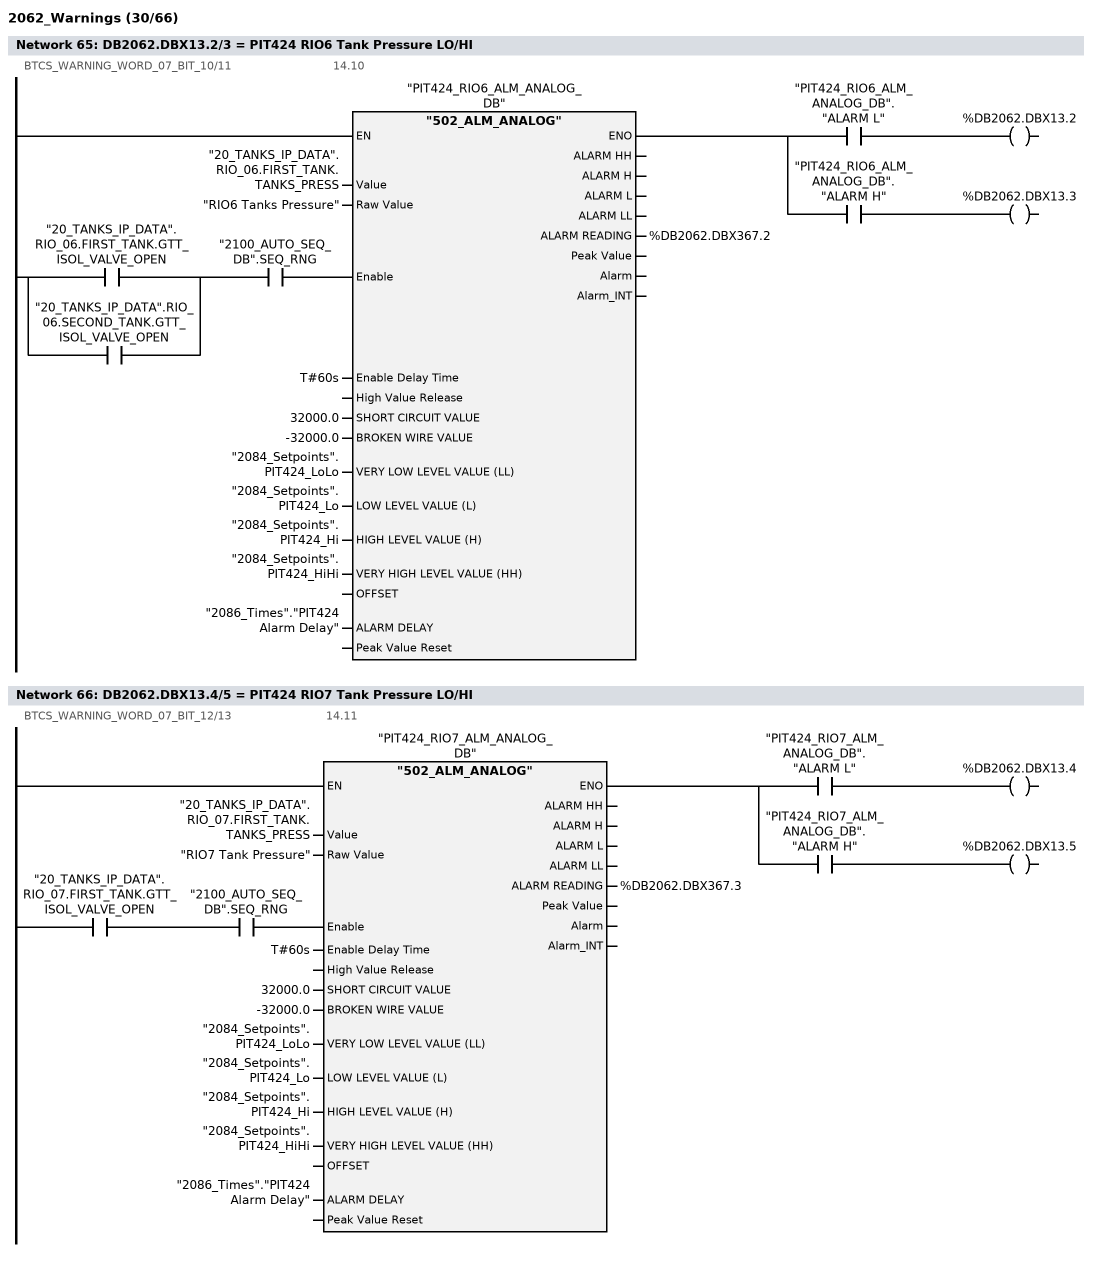
   RUNG wire#powerrail
      "PIT424_RIO6_ALM_ANALOG_DB"(Enable := wire#w2, Value := "20_TANKS_IP_DATA".RIO_06.FIRST_TANK.TANKS_PRESS, "Raw Value" := "RIO6 Tanks Pressure", "Enable Delay Time" := T#60s, "High Value Release" :=, "SHORT CIRCUIT VALUE" := 32000.0, "BROKEN WIRE VALUE" := -32000.0, "VERY LOW LEVEL VALUE (LL)" := "2084_Setpoints".PIT424_LoLo, "LOW LEVEL VALUE (L)" := "2084_Setpoints".PIT424_Lo, "HIGH LEVEL VALUE (H)" := "2084_Setpoints".PIT424_Hi, "VERY HIGH LEVEL VALUE (HH)" := "2084_Setpoints".PIT424_HiHi, OFFSET :=, "ALARM DELAY" := "2086_Times"."PIT424 Alarm Delay", "Peak Value Reset" :=, "ALARM HH" =>, "ALARM H" =>, "ALARM L" =>, "ALARM LL" =>, "ALARM READING" => %DB2062.DBX367.2, "Peak Value" =>, Alarm =>, Alarm_INT =>)
      wire#w3
      Contact( "PIT424_RIO6_ALM_ANALOG_DB"."ALARM L" )
      Coil( %DB2062.DBX13.2 )
   END_RUNG
   RUNG wire#powerrail
      Contact( "20_TANKS_IP_DATA".RIO_06.FIRST_TANK.GTT_ISOL_VALVE_OPEN )
      wire#w1
      Contact( "2100_AUTO_SEQ_DB".SEQ_RNG )
   END_RUNG wire#w2
   RUNG wire#powerrail
      Contact( "20_TANKS_IP_DATA".RIO_06.SECOND_TANK.GTT_ISOL_VALVE_OPEN )
   END_RUNG wire#w1
   RUNG wire#w3
      Contact( "PIT424_RIO6_ALM_ANALOG_DB"."ALARM H" )
      Coil( %DB2062.DBX13.3 )
   END_RUNG
   // the same network as SCL:
   "PIT424_RIO6_ALM_ANALOG_DB"(Value := "20_TANKS_IP_DATA".RIO_06.FIRST_TANK.TANKS_PRESS,   // "502_ALM_ANALOG"
                           "Raw Value" := "RIO6 Tanks Pressure",
                           Enable := ("20_TANKS_IP_DATA".RIO_06.FIRST_TANK.GTT_ISOL_VALVE_OPEN OR "20_TANKS_IP_DATA".RIO_06.SECOND_TANK.GTT_ISOL_VALVE_OPEN) AND "2100_AUTO_SEQ_DB".SEQ_RNG,
                           "Enable Delay Time" := T#60s,
                           "SHORT CIRCUIT VALUE" := 32000.0,
                           "BROKEN WIRE VALUE" := -32000.0,
                           "VERY LOW LEVEL VALUE (LL)" := "2084_Setpoints".PIT424_LoLo,
                           "LOW LEVEL VALUE (L)" := "2084_Setpoints".PIT424_Lo,
                           "HIGH LEVEL VALUE (H)" := "2084_Setpoints".PIT424_Hi,
                           "VERY HIGH LEVEL VALUE (HH)" := "2084_Setpoints".PIT424_HiHi,
                           "ALARM DELAY" := "2086_Times"."PIT424 Alarm Delay",
                           "ALARM READING" => %DB2062.DBX367.2,
                           ENO => #_w1);
   %DB2062.DBX13.2 := #_w1 AND "PIT424_RIO6_ALM_ANALOG_DB"."ALARM L";
   %DB2062.DBX13.3 := #_w1 AND "PIT424_RIO6_ALM_ANALOG_DB"."ALARM H";
END_REGION

REGION Network 66: DB2062.DBX13.4/5 = PIT424 RIO7 Tank Pressure LO/HI
   // BTCS_WARNING_WORD_07_BIT_12/13                           14.11
   RUNG wire#powerrail
      "PIT424_RIO7_ALM_ANALOG_DB"(Enable := wire#w1, Value := "20_TANKS_IP_DATA".RIO_07.FIRST_TANK.TANKS_PRESS, "Raw Value" := "RIO7 Tank Pressure", "Enable Delay Time" := T#60s, "High Value Release" :=, "SHORT CIRCUIT VALUE" := 32000.0, "BROKEN WIRE VALUE" := -32000.0, "VERY LOW LEVEL VALUE (LL)" := "2084_Setpoints".PIT424_LoLo, "LOW LEVEL VALUE (L)" := "2084_Setpoints".PIT424_Lo, "HIGH LEVEL VALUE (H)" := "2084_Setpoints".PIT424_Hi, "VERY HIGH LEVEL VALUE (HH)" := "2084_Setpoints".PIT424_HiHi, OFFSET :=, "ALARM DELAY" := "2086_Times"."PIT424 Alarm Delay", "Peak Value Reset" :=, "ALARM HH" =>, "ALARM H" =>, "ALARM L" =>, "ALARM LL" =>, "ALARM READING" => %DB2062.DBX367.3, "Peak Value" =>, Alarm =>, Alarm_INT =>)
      wire#w2
      Contact( "PIT424_RIO7_ALM_ANALOG_DB"."ALARM L" )
      Coil( %DB2062.DBX13.4 )
   END_RUNG
   RUNG wire#powerrail
      Contact( "20_TANKS_IP_DATA".RIO_07.FIRST_TANK.GTT_ISOL_VALVE_OPEN )
      Contact( "2100_AUTO_SEQ_DB".SEQ_RNG )
   END_RUNG wire#w1
   RUNG wire#w2
      Contact( "PIT424_RIO7_ALM_ANALOG_DB"."ALARM H" )
      Coil( %DB2062.DBX13.5 )
   END_RUNG
   // the same network as SCL:
   "PIT424_RIO7_ALM_ANALOG_DB"(Value := "20_TANKS_IP_DATA".RIO_07.FIRST_TANK.TANKS_PRESS,   // "502_ALM_ANALOG"
                           "Raw Value" := "RIO7 Tank Pressure",
                           Enable := "20_TANKS_IP_DATA".RIO_07.FIRST_TANK.GTT_ISOL_VALVE_OPEN AND "2100_AUTO_SEQ_DB".SEQ_RNG,
                           "Enable Delay Time" := T#60s,
                           "SHORT CIRCUIT VALUE" := 32000.0,
                           "BROKEN WIRE VALUE" := -32000.0,
                           "VERY LOW LEVEL VALUE (LL)" := "2084_Setpoints".PIT424_LoLo,
                           "LOW LEVEL VALUE (L)" := "2084_Setpoints".PIT424_Lo,
                           "HIGH LEVEL VALUE (H)" := "2084_Setpoints".PIT424_Hi,
                           "VERY HIGH LEVEL VALUE (HH)" := "2084_Setpoints".PIT424_HiHi,
                           "ALARM DELAY" := "2086_Times"."PIT424 Alarm Delay",
                           "ALARM READING" => %DB2062.DBX367.3,
                           ENO => #_w1);
   %DB2062.DBX13.4 := #_w1 AND "PIT424_RIO7_ALM_ANALOG_DB"."ALARM L";
   %DB2062.DBX13.5 := #_w1 AND "PIT424_RIO7_ALM_ANALOG_DB"."ALARM H";
END_REGION

REGION Network 67: DB2062.DBX2.6 = PIT424 Starboard Tank Pressure LO
   // BTCS_WARNING_WORD_02_BIT_6
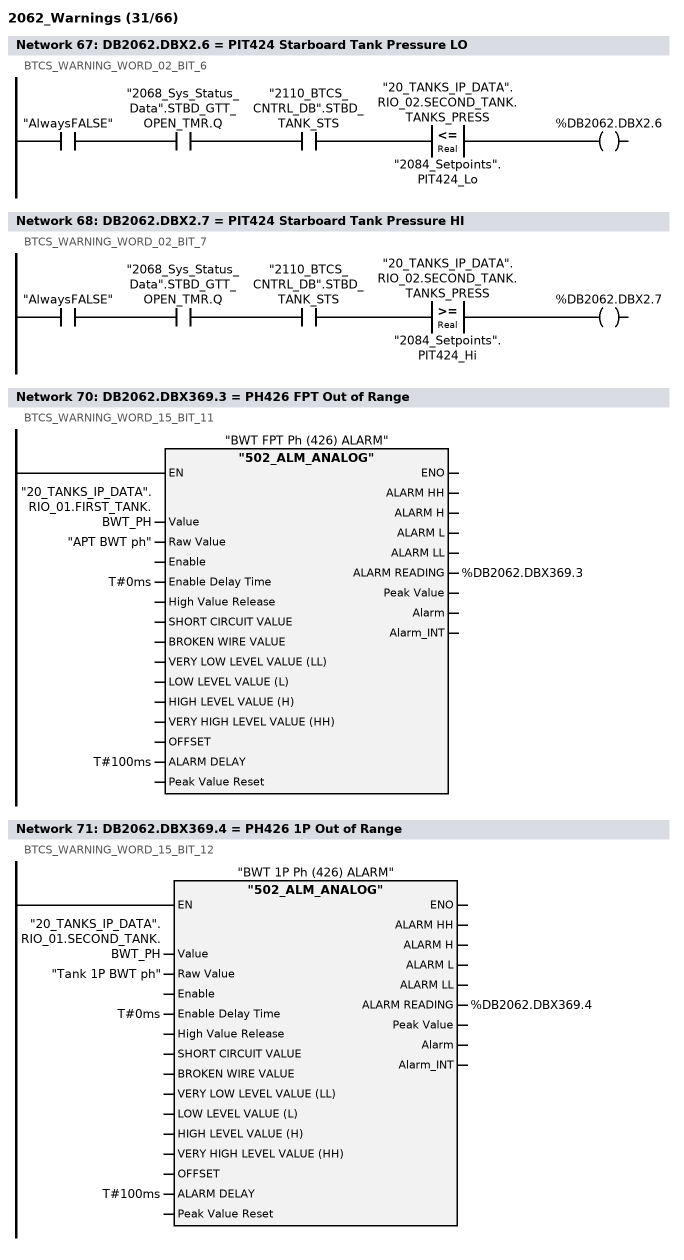
   RUNG wire#powerrail
      Contact( "AlwaysFALSE" )
      Contact( "2068_Sys_Status_Data".STBD_GTT_OPEN_TMR.Q )
      Contact( "2110_BTCS_CNTRL_DB".STBD_TANK_STS )
      { S7_Templates := "SrcType := Real" } LE_Contact(in1 := "20_TANKS_IP_DATA".RIO_02.SECOND_TANK.TANKS_PRESS, in2 := "2084_Setpoints".PIT424_Lo)
      Coil( %DB2062.DBX2.6 )
   END_RUNG
   // the same network as SCL:
   %DB2062.DBX2.6 := "AlwaysFALSE" AND "2068_Sys_Status_Data".STBD_GTT_OPEN_TMR.Q AND "2110_BTCS_CNTRL_DB".STBD_TANK_STS AND ("20_TANKS_IP_DATA".RIO_02.SECOND_TANK.TANKS_PRESS <= "2084_Setpoints".PIT424_Lo);
END_REGION

REGION Network 68: DB2062.DBX2.7 = PIT424 Starboard Tank Pressure HI
   // BTCS_WARNING_WORD_02_BIT_7
   RUNG wire#powerrail
      Contact( "AlwaysFALSE" )
      Contact( "2068_Sys_Status_Data".STBD_GTT_OPEN_TMR.Q )
      Contact( "2110_BTCS_CNTRL_DB".STBD_TANK_STS )
      { S7_Templates := "SrcType := Real" } GE_Contact(in1 := "20_TANKS_IP_DATA".RIO_02.SECOND_TANK.TANKS_PRESS, in2 := "2084_Setpoints".PIT424_Hi)
      Coil( %DB2062.DBX2.7 )
   END_RUNG
   // the same network as SCL:
   %DB2062.DBX2.7 := "AlwaysFALSE" AND "2068_Sys_Status_Data".STBD_GTT_OPEN_TMR.Q AND "2110_BTCS_CNTRL_DB".STBD_TANK_STS AND ("20_TANKS_IP_DATA".RIO_02.SECOND_TANK.TANKS_PRESS >= "2084_Setpoints".PIT424_Hi);
END_REGION

REGION Network 70: DB2062.DBX369.3 = PH426 FPT Out of Range
   // BTCS_WARNING_WORD_15_BIT_11
   RUNG wire#powerrail
      "BWT FPT Ph (426) ALARM"(Value := "20_TANKS_IP_DATA".RIO_01.FIRST_TANK.BWT_PH, "Raw Value" := "APT BWT ph", Enable :=, "Enable Delay Time" := T#0ms, "High Value Release" :=, "SHORT CIRCUIT VALUE" :=, "BROKEN WIRE VALUE" :=, "VERY LOW LEVEL VALUE (LL)" :=, "LOW LEVEL VALUE (L)" :=, "HIGH LEVEL VALUE (H)" :=, "VERY HIGH LEVEL VALUE (HH)" :=, OFFSET :=, "ALARM DELAY" := T#100ms, "Peak Value Reset" :=, "ALARM HH" =>, "ALARM H" =>, "ALARM L" =>, "ALARM LL" =>, "ALARM READING" => %DB2062.DBX369.3, "Peak Value" =>, Alarm =>, Alarm_INT =>)
   END_RUNG
   // the same network as SCL:
   "BWT FPT Ph (426) ALARM"(Value := "20_TANKS_IP_DATA".RIO_01.FIRST_TANK.BWT_PH,   // "502_ALM_ANALOG"
                           "Raw Value" := "APT BWT ph",
                           "Enable Delay Time" := T#0ms,
                           "ALARM DELAY" := T#100ms,
                           "ALARM READING" => %DB2062.DBX369.3);
END_REGION

REGION Network 71: DB2062.DBX369.4 = PH426 1P Out of Range
   // BTCS_WARNING_WORD_15_BIT_12
   RUNG wire#powerrail
      "BWT 1P Ph (426) ALARM"(Value := "20_TANKS_IP_DATA".RIO_01.SECOND_TANK.BWT_PH, "Raw Value" := "Tank 1P BWT ph", Enable :=, "Enable Delay Time" := T#0ms, "High Value Release" :=, "SHORT CIRCUIT VALUE" :=, "BROKEN WIRE VALUE" :=, "VERY LOW LEVEL VALUE (LL)" :=, "LOW LEVEL VALUE (L)" :=, "HIGH LEVEL VALUE (H)" :=, "VERY HIGH LEVEL VALUE (HH)" :=, OFFSET :=, "ALARM DELAY" := T#100ms, "Peak Value Reset" :=, "ALARM HH" =>, "ALARM H" =>, "ALARM L" =>, "ALARM LL" =>, "ALARM READING" => %DB2062.DBX369.4, "Peak Value" =>, Alarm =>, Alarm_INT =>)
   END_RUNG
   // the same network as SCL:
   "BWT 1P Ph (426) ALARM"(Value := "20_TANKS_IP_DATA".RIO_01.SECOND_TANK.BWT_PH,   // "502_ALM_ANALOG"
                           "Raw Value" := "Tank 1P BWT ph",
                           "Enable Delay Time" := T#0ms,
                           "ALARM DELAY" := T#100ms,
                           "ALARM READING" => %DB2062.DBX369.4);
END_REGION

REGION Network 72: DB2062.DBX369.5 = PH425 1S Out of Range
   // BTCS_WARNING_WORD_15_BIT_13
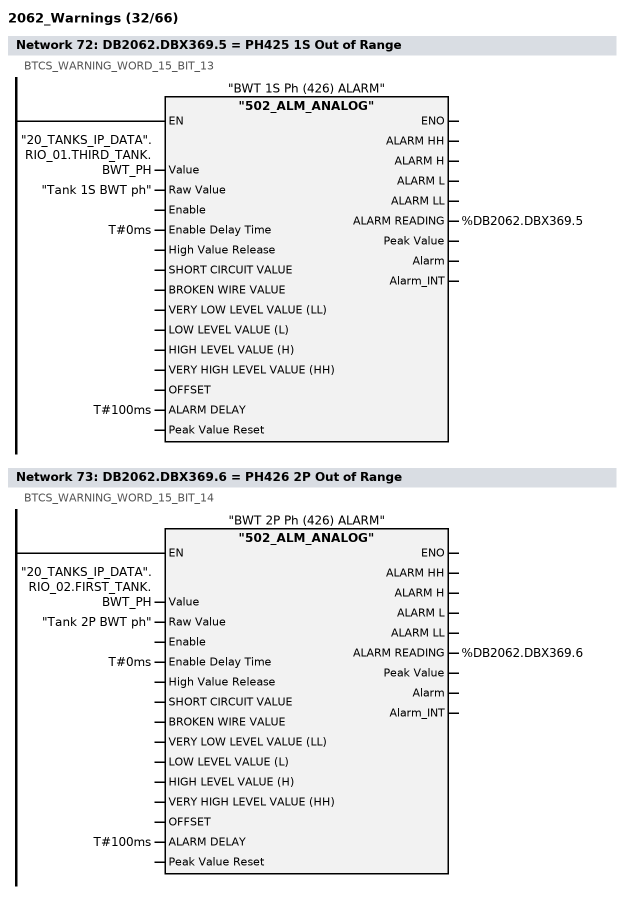
   RUNG wire#powerrail
      "BWT 1S Ph (426) ALARM"(Value := "20_TANKS_IP_DATA".RIO_01.THIRD_TANK.BWT_PH, "Raw Value" := "Tank 1S BWT ph", Enable :=, "Enable Delay Time" := T#0ms, "High Value Release" :=, "SHORT CIRCUIT VALUE" :=, "BROKEN WIRE VALUE" :=, "VERY LOW LEVEL VALUE (LL)" :=, "LOW LEVEL VALUE (L)" :=, "HIGH LEVEL VALUE (H)" :=, "VERY HIGH LEVEL VALUE (HH)" :=, OFFSET :=, "ALARM DELAY" := T#100ms, "Peak Value Reset" :=, "ALARM HH" =>, "ALARM H" =>, "ALARM L" =>, "ALARM LL" =>, "ALARM READING" => %DB2062.DBX369.5, "Peak Value" =>, Alarm =>, Alarm_INT =>)
   END_RUNG
   // the same network as SCL:
   "BWT 1S Ph (426) ALARM"(Value := "20_TANKS_IP_DATA".RIO_01.THIRD_TANK.BWT_PH,   // "502_ALM_ANALOG"
                           "Raw Value" := "Tank 1S BWT ph",
                           "Enable Delay Time" := T#0ms,
                           "ALARM DELAY" := T#100ms,
                           "ALARM READING" => %DB2062.DBX369.5);
END_REGION

REGION Network 73: DB2062.DBX369.6 = PH426 2P Out of Range
   // BTCS_WARNING_WORD_15_BIT_14
   RUNG wire#powerrail
      "BWT 2P Ph (426) ALARM"(Value := "20_TANKS_IP_DATA".RIO_02.FIRST_TANK.BWT_PH, "Raw Value" := "Tank 2P BWT ph", Enable :=, "Enable Delay Time" := T#0ms, "High Value Release" :=, "SHORT CIRCUIT VALUE" :=, "BROKEN WIRE VALUE" :=, "VERY LOW LEVEL VALUE (LL)" :=, "LOW LEVEL VALUE (L)" :=, "HIGH LEVEL VALUE (H)" :=, "VERY HIGH LEVEL VALUE (HH)" :=, OFFSET :=, "ALARM DELAY" := T#100ms, "Peak Value Reset" :=, "ALARM HH" =>, "ALARM H" =>, "ALARM L" =>, "ALARM LL" =>, "ALARM READING" => %DB2062.DBX369.6, "Peak Value" =>, Alarm =>, Alarm_INT =>)
   END_RUNG
   // the same network as SCL:
   "BWT 2P Ph (426) ALARM"(Value := "20_TANKS_IP_DATA".RIO_02.FIRST_TANK.BWT_PH,   // "502_ALM_ANALOG"
                           "Raw Value" := "Tank 2P BWT ph",
                           "Enable Delay Time" := T#0ms,
                           "ALARM DELAY" := T#100ms,
                           "ALARM READING" => %DB2062.DBX369.6);
END_REGION

REGION Network 74: DB2062.DBX369.7 = PH425 2S Out of Range
   // BTCS_WARNING_WORD_15_BIT_15
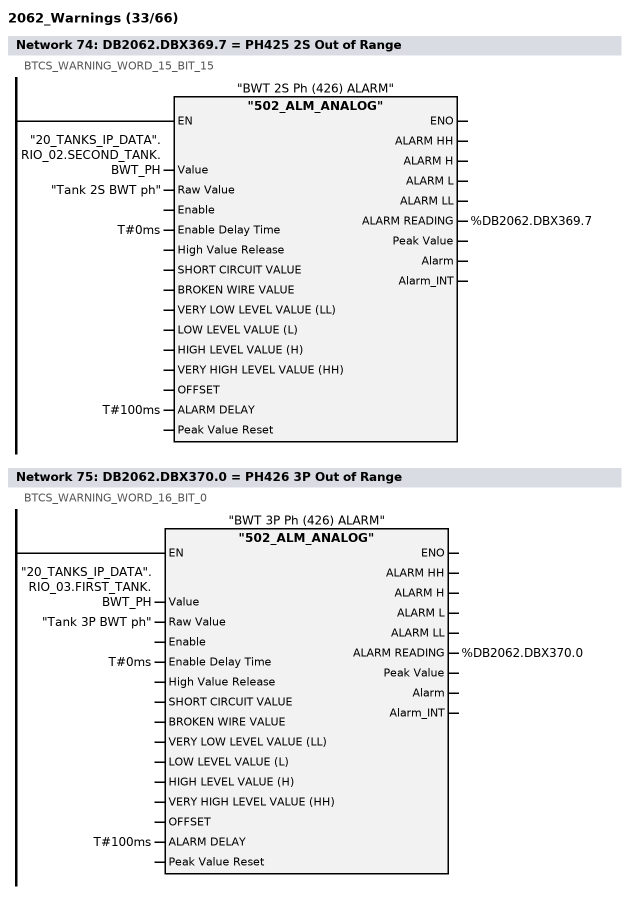
   RUNG wire#powerrail
      "BWT 2S Ph (426) ALARM"(Value := "20_TANKS_IP_DATA".RIO_02.SECOND_TANK.BWT_PH, "Raw Value" := "Tank 2S BWT ph", Enable :=, "Enable Delay Time" := T#0ms, "High Value Release" :=, "SHORT CIRCUIT VALUE" :=, "BROKEN WIRE VALUE" :=, "VERY LOW LEVEL VALUE (LL)" :=, "LOW LEVEL VALUE (L)" :=, "HIGH LEVEL VALUE (H)" :=, "VERY HIGH LEVEL VALUE (HH)" :=, OFFSET :=, "ALARM DELAY" := T#100ms, "Peak Value Reset" :=, "ALARM HH" =>, "ALARM H" =>, "ALARM L" =>, "ALARM LL" =>, "ALARM READING" => %DB2062.DBX369.7, "Peak Value" =>, Alarm =>, Alarm_INT =>)
   END_RUNG
   // the same network as SCL:
   "BWT 2S Ph (426) ALARM"(Value := "20_TANKS_IP_DATA".RIO_02.SECOND_TANK.BWT_PH,   // "502_ALM_ANALOG"
                           "Raw Value" := "Tank 2S BWT ph",
                           "Enable Delay Time" := T#0ms,
                           "ALARM DELAY" := T#100ms,
                           "ALARM READING" => %DB2062.DBX369.7);
END_REGION

REGION Network 75: DB2062.DBX370.0 = PH426 3P Out of Range
   // BTCS_WARNING_WORD_16_BIT_0
   RUNG wire#powerrail
      "BWT 3P Ph (426) ALARM"(Value := "20_TANKS_IP_DATA".RIO_03.FIRST_TANK.BWT_PH, "Raw Value" := "Tank 3P BWT ph", Enable :=, "Enable Delay Time" := T#0ms, "High Value Release" :=, "SHORT CIRCUIT VALUE" :=, "BROKEN WIRE VALUE" :=, "VERY LOW LEVEL VALUE (LL)" :=, "LOW LEVEL VALUE (L)" :=, "HIGH LEVEL VALUE (H)" :=, "VERY HIGH LEVEL VALUE (HH)" :=, OFFSET :=, "ALARM DELAY" := T#100ms, "Peak Value Reset" :=, "ALARM HH" =>, "ALARM H" =>, "ALARM L" =>, "ALARM LL" =>, "ALARM READING" => %DB2062.DBX370.0, "Peak Value" =>, Alarm =>, Alarm_INT =>)
   END_RUNG
   // the same network as SCL:
   "BWT 3P Ph (426) ALARM"(Value := "20_TANKS_IP_DATA".RIO_03.FIRST_TANK.BWT_PH,   // "502_ALM_ANALOG"
                           "Raw Value" := "Tank 3P BWT ph",
                           "Enable Delay Time" := T#0ms,
                           "ALARM DELAY" := T#100ms,
                           "ALARM READING" => %DB2062.DBX370.0);
END_REGION

REGION Network 76: DB2062.DBX370.1 = PH425 3S Out of Range
   // BTCS_WARNING_WORD_16_BIT_1
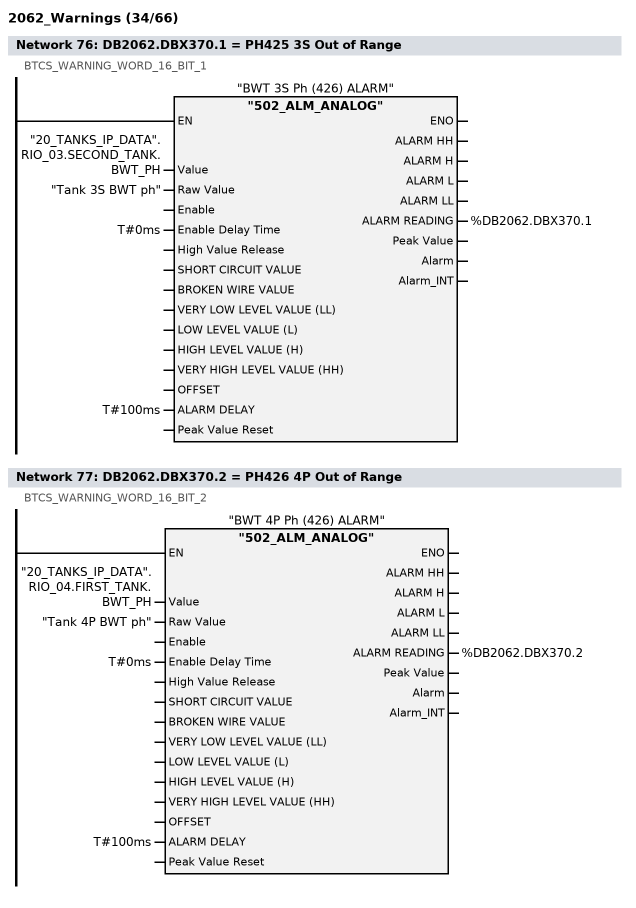
   RUNG wire#powerrail
      "BWT 3S Ph (426) ALARM"(Value := "20_TANKS_IP_DATA".RIO_03.SECOND_TANK.BWT_PH, "Raw Value" := "Tank 3S BWT ph", Enable :=, "Enable Delay Time" := T#0ms, "High Value Release" :=, "SHORT CIRCUIT VALUE" :=, "BROKEN WIRE VALUE" :=, "VERY LOW LEVEL VALUE (LL)" :=, "LOW LEVEL VALUE (L)" :=, "HIGH LEVEL VALUE (H)" :=, "VERY HIGH LEVEL VALUE (HH)" :=, OFFSET :=, "ALARM DELAY" := T#100ms, "Peak Value Reset" :=, "ALARM HH" =>, "ALARM H" =>, "ALARM L" =>, "ALARM LL" =>, "ALARM READING" => %DB2062.DBX370.1, "Peak Value" =>, Alarm =>, Alarm_INT =>)
   END_RUNG
   // the same network as SCL:
   "BWT 3S Ph (426) ALARM"(Value := "20_TANKS_IP_DATA".RIO_03.SECOND_TANK.BWT_PH,   // "502_ALM_ANALOG"
                           "Raw Value" := "Tank 3S BWT ph",
                           "Enable Delay Time" := T#0ms,
                           "ALARM DELAY" := T#100ms,
                           "ALARM READING" => %DB2062.DBX370.1);
END_REGION

REGION Network 77: DB2062.DBX370.2 = PH426 4P Out of Range
   // BTCS_WARNING_WORD_16_BIT_2
   RUNG wire#powerrail
      "BWT 4P Ph (426) ALARM"(Value := "20_TANKS_IP_DATA".RIO_04.FIRST_TANK.BWT_PH, "Raw Value" := "Tank 4P BWT ph", Enable :=, "Enable Delay Time" := T#0ms, "High Value Release" :=, "SHORT CIRCUIT VALUE" :=, "BROKEN WIRE VALUE" :=, "VERY LOW LEVEL VALUE (LL)" :=, "LOW LEVEL VALUE (L)" :=, "HIGH LEVEL VALUE (H)" :=, "VERY HIGH LEVEL VALUE (HH)" :=, OFFSET :=, "ALARM DELAY" := T#100ms, "Peak Value Reset" :=, "ALARM HH" =>, "ALARM H" =>, "ALARM L" =>, "ALARM LL" =>, "ALARM READING" => %DB2062.DBX370.2, "Peak Value" =>, Alarm =>, Alarm_INT =>)
   END_RUNG
   // the same network as SCL:
   "BWT 4P Ph (426) ALARM"(Value := "20_TANKS_IP_DATA".RIO_04.FIRST_TANK.BWT_PH,   // "502_ALM_ANALOG"
                           "Raw Value" := "Tank 4P BWT ph",
                           "Enable Delay Time" := T#0ms,
                           "ALARM DELAY" := T#100ms,
                           "ALARM READING" => %DB2062.DBX370.2);
END_REGION

REGION Network 78: DB2062.DBX370.4 = PH425 4S Out of Range
   // BTCS_WARNING_WORD_16_BIT_4
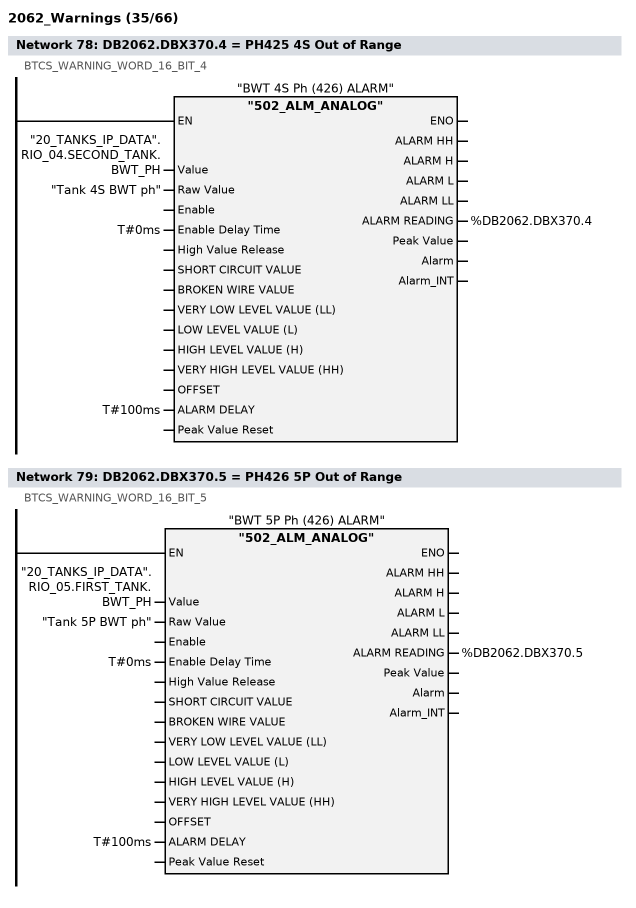
   RUNG wire#powerrail
      "BWT 4S Ph (426) ALARM"(Value := "20_TANKS_IP_DATA".RIO_04.SECOND_TANK.BWT_PH, "Raw Value" := "Tank 4S BWT ph", Enable :=, "Enable Delay Time" := T#0ms, "High Value Release" :=, "SHORT CIRCUIT VALUE" :=, "BROKEN WIRE VALUE" :=, "VERY LOW LEVEL VALUE (LL)" :=, "LOW LEVEL VALUE (L)" :=, "HIGH LEVEL VALUE (H)" :=, "VERY HIGH LEVEL VALUE (HH)" :=, OFFSET :=, "ALARM DELAY" := T#100ms, "Peak Value Reset" :=, "ALARM HH" =>, "ALARM H" =>, "ALARM L" =>, "ALARM LL" =>, "ALARM READING" => %DB2062.DBX370.4, "Peak Value" =>, Alarm =>, Alarm_INT =>)
   END_RUNG
   // the same network as SCL:
   "BWT 4S Ph (426) ALARM"(Value := "20_TANKS_IP_DATA".RIO_04.SECOND_TANK.BWT_PH,   // "502_ALM_ANALOG"
                           "Raw Value" := "Tank 4S BWT ph",
                           "Enable Delay Time" := T#0ms,
                           "ALARM DELAY" := T#100ms,
                           "ALARM READING" => %DB2062.DBX370.4);
END_REGION

REGION Network 79: DB2062.DBX370.5 = PH426 5P Out of Range
   // BTCS_WARNING_WORD_16_BIT_5
   RUNG wire#powerrail
      "BWT 5P Ph (426) ALARM"(Value := "20_TANKS_IP_DATA".RIO_05.FIRST_TANK.BWT_PH, "Raw Value" := "Tank 5P BWT ph", Enable :=, "Enable Delay Time" := T#0ms, "High Value Release" :=, "SHORT CIRCUIT VALUE" :=, "BROKEN WIRE VALUE" :=, "VERY LOW LEVEL VALUE (LL)" :=, "LOW LEVEL VALUE (L)" :=, "HIGH LEVEL VALUE (H)" :=, "VERY HIGH LEVEL VALUE (HH)" :=, OFFSET :=, "ALARM DELAY" := T#100ms, "Peak Value Reset" :=, "ALARM HH" =>, "ALARM H" =>, "ALARM L" =>, "ALARM LL" =>, "ALARM READING" => %DB2062.DBX370.5, "Peak Value" =>, Alarm =>, Alarm_INT =>)
   END_RUNG
   // the same network as SCL:
   "BWT 5P Ph (426) ALARM"(Value := "20_TANKS_IP_DATA".RIO_05.FIRST_TANK.BWT_PH,   // "502_ALM_ANALOG"
                           "Raw Value" := "Tank 5P BWT ph",
                           "Enable Delay Time" := T#0ms,
                           "ALARM DELAY" := T#100ms,
                           "ALARM READING" => %DB2062.DBX370.5);
END_REGION

REGION Network 80: DB2062.DBX370.6 = PH425 5S Out of Range
   // BTCS_WARNING_WORD_16_BIT_6
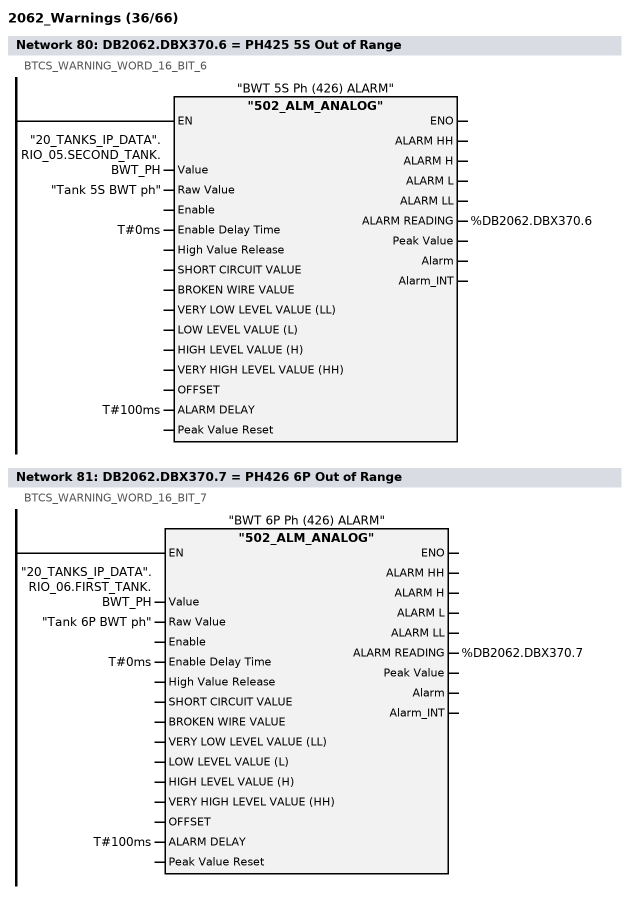
   RUNG wire#powerrail
      "BWT 5S Ph (426) ALARM"(Value := "20_TANKS_IP_DATA".RIO_05.SECOND_TANK.BWT_PH, "Raw Value" := "Tank 5S BWT ph", Enable :=, "Enable Delay Time" := T#0ms, "High Value Release" :=, "SHORT CIRCUIT VALUE" :=, "BROKEN WIRE VALUE" :=, "VERY LOW LEVEL VALUE (LL)" :=, "LOW LEVEL VALUE (L)" :=, "HIGH LEVEL VALUE (H)" :=, "VERY HIGH LEVEL VALUE (HH)" :=, OFFSET :=, "ALARM DELAY" := T#100ms, "Peak Value Reset" :=, "ALARM HH" =>, "ALARM H" =>, "ALARM L" =>, "ALARM LL" =>, "ALARM READING" => %DB2062.DBX370.6, "Peak Value" =>, Alarm =>, Alarm_INT =>)
   END_RUNG
   // the same network as SCL:
   "BWT 5S Ph (426) ALARM"(Value := "20_TANKS_IP_DATA".RIO_05.SECOND_TANK.BWT_PH,   // "502_ALM_ANALOG"
                           "Raw Value" := "Tank 5S BWT ph",
                           "Enable Delay Time" := T#0ms,
                           "ALARM DELAY" := T#100ms,
                           "ALARM READING" => %DB2062.DBX370.6);
END_REGION

REGION Network 81: DB2062.DBX370.7 = PH426 6P Out of Range
   // BTCS_WARNING_WORD_16_BIT_7
   RUNG wire#powerrail
      "BWT 6P Ph (426) ALARM"(Value := "20_TANKS_IP_DATA".RIO_06.FIRST_TANK.BWT_PH, "Raw Value" := "Tank 6P BWT ph", Enable :=, "Enable Delay Time" := T#0ms, "High Value Release" :=, "SHORT CIRCUIT VALUE" :=, "BROKEN WIRE VALUE" :=, "VERY LOW LEVEL VALUE (LL)" :=, "LOW LEVEL VALUE (L)" :=, "HIGH LEVEL VALUE (H)" :=, "VERY HIGH LEVEL VALUE (HH)" :=, OFFSET :=, "ALARM DELAY" := T#100ms, "Peak Value Reset" :=, "ALARM HH" =>, "ALARM H" =>, "ALARM L" =>, "ALARM LL" =>, "ALARM READING" => %DB2062.DBX370.7, "Peak Value" =>, Alarm =>, Alarm_INT =>)
   END_RUNG
   // the same network as SCL:
   "BWT 6P Ph (426) ALARM"(Value := "20_TANKS_IP_DATA".RIO_06.FIRST_TANK.BWT_PH,   // "502_ALM_ANALOG"
                           "Raw Value" := "Tank 6P BWT ph",
                           "Enable Delay Time" := T#0ms,
                           "ALARM DELAY" := T#100ms,
                           "ALARM READING" => %DB2062.DBX370.7);
END_REGION

REGION Network 82: DB2062.DBX371.0 = PH425 6S Out of Range
   // BTCS_WARNING_WORD_16_BIT_8
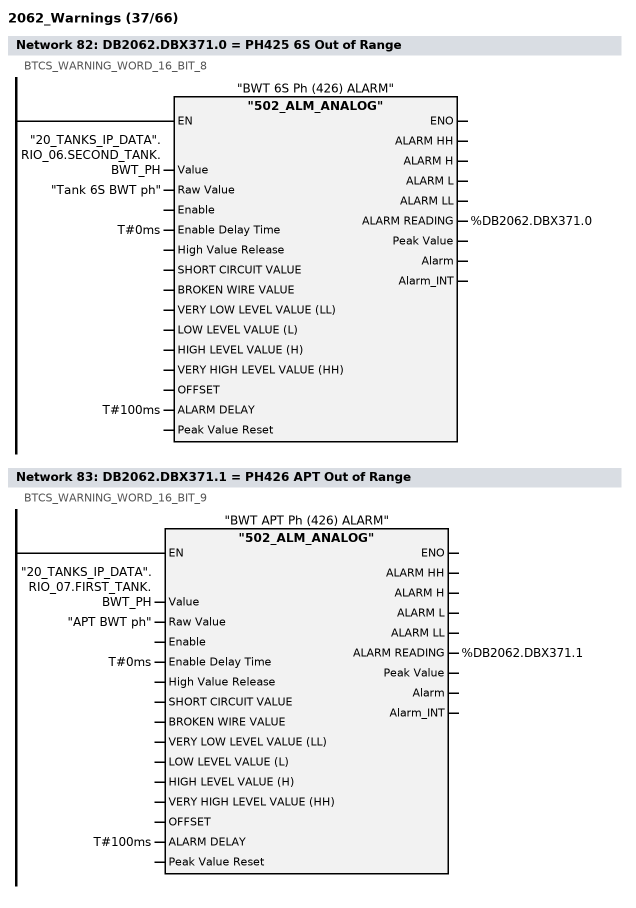
   RUNG wire#powerrail
      "BWT 6S Ph (426) ALARM"(Value := "20_TANKS_IP_DATA".RIO_06.SECOND_TANK.BWT_PH, "Raw Value" := "Tank 6S BWT ph", Enable :=, "Enable Delay Time" := T#0ms, "High Value Release" :=, "SHORT CIRCUIT VALUE" :=, "BROKEN WIRE VALUE" :=, "VERY LOW LEVEL VALUE (LL)" :=, "LOW LEVEL VALUE (L)" :=, "HIGH LEVEL VALUE (H)" :=, "VERY HIGH LEVEL VALUE (HH)" :=, OFFSET :=, "ALARM DELAY" := T#100ms, "Peak Value Reset" :=, "ALARM HH" =>, "ALARM H" =>, "ALARM L" =>, "ALARM LL" =>, "ALARM READING" => %DB2062.DBX371.0, "Peak Value" =>, Alarm =>, Alarm_INT =>)
   END_RUNG
   // the same network as SCL:
   "BWT 6S Ph (426) ALARM"(Value := "20_TANKS_IP_DATA".RIO_06.SECOND_TANK.BWT_PH,   // "502_ALM_ANALOG"
                           "Raw Value" := "Tank 6S BWT ph",
                           "Enable Delay Time" := T#0ms,
                           "ALARM DELAY" := T#100ms,
                           "ALARM READING" => %DB2062.DBX371.0);
END_REGION

REGION Network 83: DB2062.DBX371.1 = PH426 APT Out of Range
   // BTCS_WARNING_WORD_16_BIT_9
   RUNG wire#powerrail
      "BWT APT Ph (426) ALARM"(Value := "20_TANKS_IP_DATA".RIO_07.FIRST_TANK.BWT_PH, "Raw Value" := "APT BWT ph", Enable :=, "Enable Delay Time" := T#0ms, "High Value Release" :=, "SHORT CIRCUIT VALUE" :=, "BROKEN WIRE VALUE" :=, "VERY LOW LEVEL VALUE (LL)" :=, "LOW LEVEL VALUE (L)" :=, "HIGH LEVEL VALUE (H)" :=, "VERY HIGH LEVEL VALUE (HH)" :=, OFFSET :=, "ALARM DELAY" := T#100ms, "Peak Value Reset" :=, "ALARM HH" =>, "ALARM H" =>, "ALARM L" =>, "ALARM LL" =>, "ALARM READING" => %DB2062.DBX371.1, "Peak Value" =>, Alarm =>, Alarm_INT =>)
   END_RUNG
   // the same network as SCL:
   "BWT APT Ph (426) ALARM"(Value := "20_TANKS_IP_DATA".RIO_07.FIRST_TANK.BWT_PH,   // "502_ALM_ANALOG"
                           "Raw Value" := "APT BWT ph",
                           "Enable Delay Time" := T#0ms,
                           "ALARM DELAY" := T#100ms,
                           "ALARM READING" => %DB2062.DBX371.1);
END_REGION

REGION Network 85: DB2062.DBX371.2 = DO426 FPT
   // BTCS_WARNING_WORD_16_BIT_10
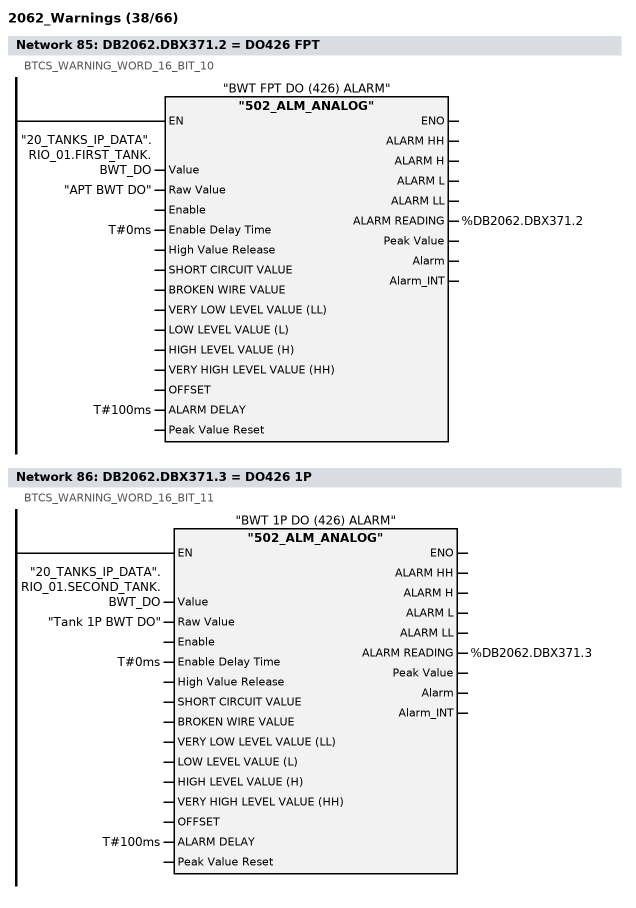
   RUNG wire#powerrail
      "BWT FPT DO (426) ALARM"(Value := "20_TANKS_IP_DATA".RIO_01.FIRST_TANK.BWT_DO, "Raw Value" := "APT BWT DO", Enable :=, "Enable Delay Time" := T#0ms, "High Value Release" :=, "SHORT CIRCUIT VALUE" :=, "BROKEN WIRE VALUE" :=, "VERY LOW LEVEL VALUE (LL)" :=, "LOW LEVEL VALUE (L)" :=, "HIGH LEVEL VALUE (H)" :=, "VERY HIGH LEVEL VALUE (HH)" :=, OFFSET :=, "ALARM DELAY" := T#100ms, "Peak Value Reset" :=, "ALARM HH" =>, "ALARM H" =>, "ALARM L" =>, "ALARM LL" =>, "ALARM READING" => %DB2062.DBX371.2, "Peak Value" =>, Alarm =>, Alarm_INT =>)
   END_RUNG
   // the same network as SCL:
   "BWT FPT DO (426) ALARM"(Value := "20_TANKS_IP_DATA".RIO_01.FIRST_TANK.BWT_DO,   // "502_ALM_ANALOG"
                           "Raw Value" := "APT BWT DO",
                           "Enable Delay Time" := T#0ms,
                           "ALARM DELAY" := T#100ms,
                           "ALARM READING" => %DB2062.DBX371.2);
END_REGION

REGION Network 86: DB2062.DBX371.3 = DO426 1P
   // BTCS_WARNING_WORD_16_BIT_11
   RUNG wire#powerrail
      "BWT 1P DO (426) ALARM"(Value := "20_TANKS_IP_DATA".RIO_01.SECOND_TANK.BWT_DO, "Raw Value" := "Tank 1P BWT DO", Enable :=, "Enable Delay Time" := T#0ms, "High Value Release" :=, "SHORT CIRCUIT VALUE" :=, "BROKEN WIRE VALUE" :=, "VERY LOW LEVEL VALUE (LL)" :=, "LOW LEVEL VALUE (L)" :=, "HIGH LEVEL VALUE (H)" :=, "VERY HIGH LEVEL VALUE (HH)" :=, OFFSET :=, "ALARM DELAY" := T#100ms, "Peak Value Reset" :=, "ALARM HH" =>, "ALARM H" =>, "ALARM L" =>, "ALARM LL" =>, "ALARM READING" => %DB2062.DBX371.3, "Peak Value" =>, Alarm =>, Alarm_INT =>)
   END_RUNG
   // the same network as SCL:
   "BWT 1P DO (426) ALARM"(Value := "20_TANKS_IP_DATA".RIO_01.SECOND_TANK.BWT_DO,   // "502_ALM_ANALOG"
                           "Raw Value" := "Tank 1P BWT DO",
                           "Enable Delay Time" := T#0ms,
                           "ALARM DELAY" := T#100ms,
                           "ALARM READING" => %DB2062.DBX371.3);
END_REGION

REGION Network 87: DB2062.DBX371.4 = DO426 1S
   // BTCS_WARNING_WORD_16_BIT_12
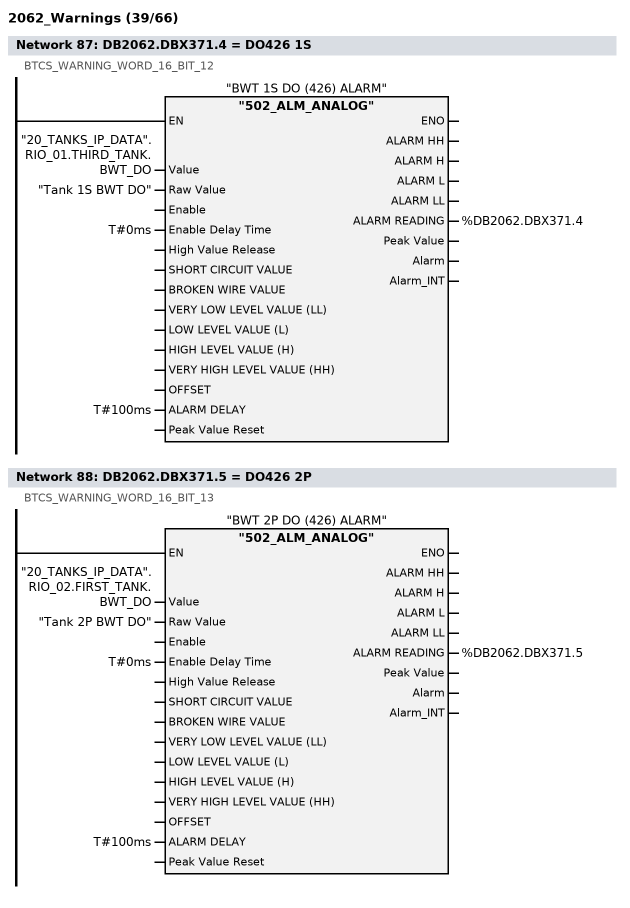
   RUNG wire#powerrail
      "BWT 1S DO (426) ALARM"(Value := "20_TANKS_IP_DATA".RIO_01.THIRD_TANK.BWT_DO, "Raw Value" := "Tank 1S BWT DO", Enable :=, "Enable Delay Time" := T#0ms, "High Value Release" :=, "SHORT CIRCUIT VALUE" :=, "BROKEN WIRE VALUE" :=, "VERY LOW LEVEL VALUE (LL)" :=, "LOW LEVEL VALUE (L)" :=, "HIGH LEVEL VALUE (H)" :=, "VERY HIGH LEVEL VALUE (HH)" :=, OFFSET :=, "ALARM DELAY" := T#100ms, "Peak Value Reset" :=, "ALARM HH" =>, "ALARM H" =>, "ALARM L" =>, "ALARM LL" =>, "ALARM READING" => %DB2062.DBX371.4, "Peak Value" =>, Alarm =>, Alarm_INT =>)
   END_RUNG
   // the same network as SCL:
   "BWT 1S DO (426) ALARM"(Value := "20_TANKS_IP_DATA".RIO_01.THIRD_TANK.BWT_DO,   // "502_ALM_ANALOG"
                           "Raw Value" := "Tank 1S BWT DO",
                           "Enable Delay Time" := T#0ms,
                           "ALARM DELAY" := T#100ms,
                           "ALARM READING" => %DB2062.DBX371.4);
END_REGION

REGION Network 88: DB2062.DBX371.5 = DO426 2P
   // BTCS_WARNING_WORD_16_BIT_13
   RUNG wire#powerrail
      "BWT 2P DO (426) ALARM"(Value := "20_TANKS_IP_DATA".RIO_02.FIRST_TANK.BWT_DO, "Raw Value" := "Tank 2P BWT DO", Enable :=, "Enable Delay Time" := T#0ms, "High Value Release" :=, "SHORT CIRCUIT VALUE" :=, "BROKEN WIRE VALUE" :=, "VERY LOW LEVEL VALUE (LL)" :=, "LOW LEVEL VALUE (L)" :=, "HIGH LEVEL VALUE (H)" :=, "VERY HIGH LEVEL VALUE (HH)" :=, OFFSET :=, "ALARM DELAY" := T#100ms, "Peak Value Reset" :=, "ALARM HH" =>, "ALARM H" =>, "ALARM L" =>, "ALARM LL" =>, "ALARM READING" => %DB2062.DBX371.5, "Peak Value" =>, Alarm =>, Alarm_INT =>)
   END_RUNG
   // the same network as SCL:
   "BWT 2P DO (426) ALARM"(Value := "20_TANKS_IP_DATA".RIO_02.FIRST_TANK.BWT_DO,   // "502_ALM_ANALOG"
                           "Raw Value" := "Tank 2P BWT DO",
                           "Enable Delay Time" := T#0ms,
                           "ALARM DELAY" := T#100ms,
                           "ALARM READING" => %DB2062.DBX371.5);
END_REGION

REGION Network 89: DB2062.DBX371.6 = DO426 2S
   // BTCS_WARNING_WORD_16_BIT_14
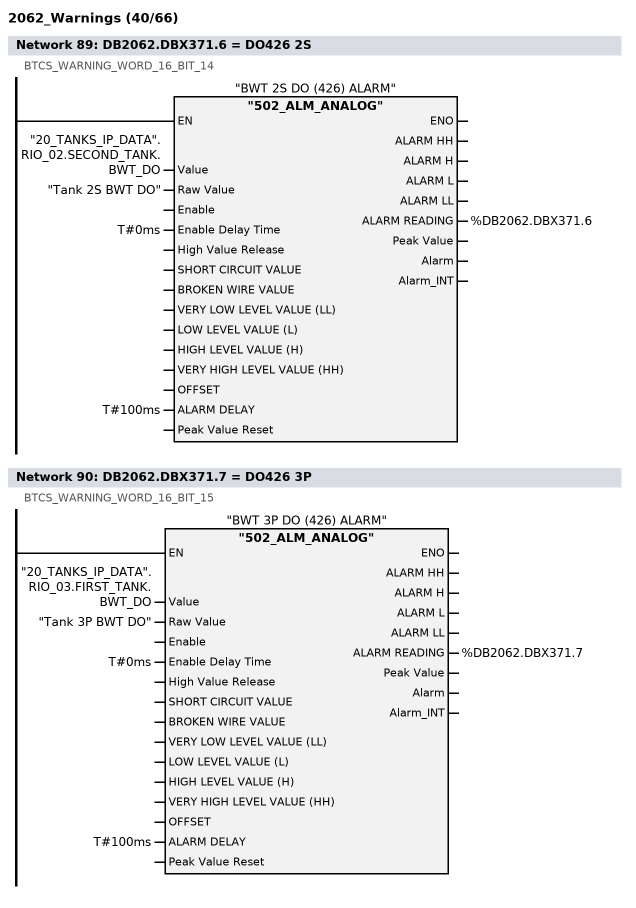
   RUNG wire#powerrail
      "BWT 2S DO (426) ALARM"(Value := "20_TANKS_IP_DATA".RIO_02.SECOND_TANK.BWT_DO, "Raw Value" := "Tank 2S BWT DO", Enable :=, "Enable Delay Time" := T#0ms, "High Value Release" :=, "SHORT CIRCUIT VALUE" :=, "BROKEN WIRE VALUE" :=, "VERY LOW LEVEL VALUE (LL)" :=, "LOW LEVEL VALUE (L)" :=, "HIGH LEVEL VALUE (H)" :=, "VERY HIGH LEVEL VALUE (HH)" :=, OFFSET :=, "ALARM DELAY" := T#100ms, "Peak Value Reset" :=, "ALARM HH" =>, "ALARM H" =>, "ALARM L" =>, "ALARM LL" =>, "ALARM READING" => %DB2062.DBX371.6, "Peak Value" =>, Alarm =>, Alarm_INT =>)
   END_RUNG
   // the same network as SCL:
   "BWT 2S DO (426) ALARM"(Value := "20_TANKS_IP_DATA".RIO_02.SECOND_TANK.BWT_DO,   // "502_ALM_ANALOG"
                           "Raw Value" := "Tank 2S BWT DO",
                           "Enable Delay Time" := T#0ms,
                           "ALARM DELAY" := T#100ms,
                           "ALARM READING" => %DB2062.DBX371.6);
END_REGION

REGION Network 90: DB2062.DBX371.7 = DO426 3P
   // BTCS_WARNING_WORD_16_BIT_15
   RUNG wire#powerrail
      "BWT 3P DO (426) ALARM"(Value := "20_TANKS_IP_DATA".RIO_03.FIRST_TANK.BWT_DO, "Raw Value" := "Tank 3P BWT DO", Enable :=, "Enable Delay Time" := T#0ms, "High Value Release" :=, "SHORT CIRCUIT VALUE" :=, "BROKEN WIRE VALUE" :=, "VERY LOW LEVEL VALUE (LL)" :=, "LOW LEVEL VALUE (L)" :=, "HIGH LEVEL VALUE (H)" :=, "VERY HIGH LEVEL VALUE (HH)" :=, OFFSET :=, "ALARM DELAY" := T#100ms, "Peak Value Reset" :=, "ALARM HH" =>, "ALARM H" =>, "ALARM L" =>, "ALARM LL" =>, "ALARM READING" => %DB2062.DBX371.7, "Peak Value" =>, Alarm =>, Alarm_INT =>)
   END_RUNG
   // the same network as SCL:
   "BWT 3P DO (426) ALARM"(Value := "20_TANKS_IP_DATA".RIO_03.FIRST_TANK.BWT_DO,   // "502_ALM_ANALOG"
                           "Raw Value" := "Tank 3P BWT DO",
                           "Enable Delay Time" := T#0ms,
                           "ALARM DELAY" := T#100ms,
                           "ALARM READING" => %DB2062.DBX371.7);
END_REGION

REGION Network 91: DB2062.DBX372.0 = DO426 3S
   // BTCS_WARNING_WORD_17_BIT_0
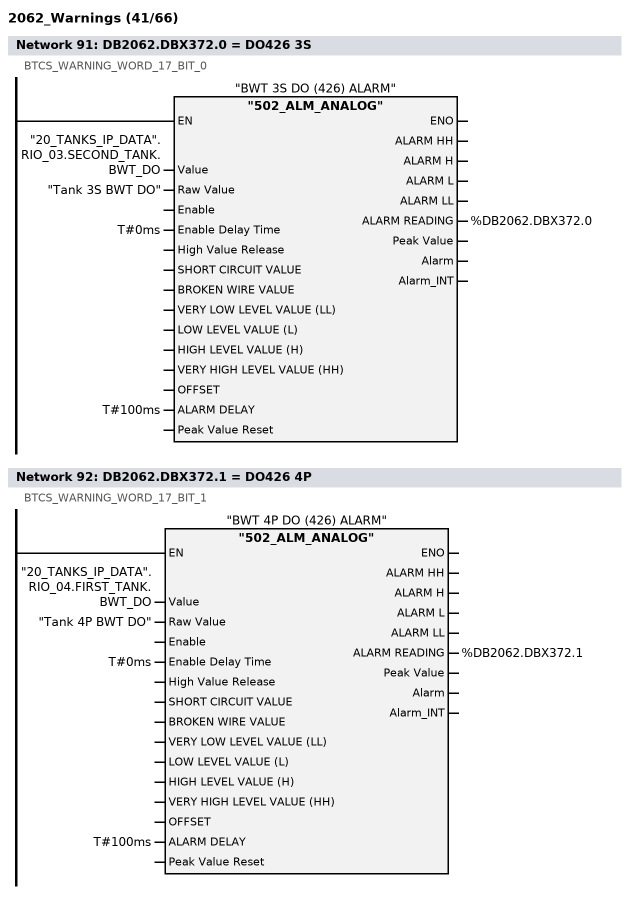
   RUNG wire#powerrail
      "BWT 3S DO (426) ALARM"(Value := "20_TANKS_IP_DATA".RIO_03.SECOND_TANK.BWT_DO, "Raw Value" := "Tank 3S BWT DO", Enable :=, "Enable Delay Time" := T#0ms, "High Value Release" :=, "SHORT CIRCUIT VALUE" :=, "BROKEN WIRE VALUE" :=, "VERY LOW LEVEL VALUE (LL)" :=, "LOW LEVEL VALUE (L)" :=, "HIGH LEVEL VALUE (H)" :=, "VERY HIGH LEVEL VALUE (HH)" :=, OFFSET :=, "ALARM DELAY" := T#100ms, "Peak Value Reset" :=, "ALARM HH" =>, "ALARM H" =>, "ALARM L" =>, "ALARM LL" =>, "ALARM READING" => %DB2062.DBX372.0, "Peak Value" =>, Alarm =>, Alarm_INT =>)
   END_RUNG
   // the same network as SCL:
   "BWT 3S DO (426) ALARM"(Value := "20_TANKS_IP_DATA".RIO_03.SECOND_TANK.BWT_DO,   // "502_ALM_ANALOG"
                           "Raw Value" := "Tank 3S BWT DO",
                           "Enable Delay Time" := T#0ms,
                           "ALARM DELAY" := T#100ms,
                           "ALARM READING" => %DB2062.DBX372.0);
END_REGION

REGION Network 92: DB2062.DBX372.1 = DO426 4P
   // BTCS_WARNING_WORD_17_BIT_1
   RUNG wire#powerrail
      "BWT 4P DO (426) ALARM"(Value := "20_TANKS_IP_DATA".RIO_04.FIRST_TANK.BWT_DO, "Raw Value" := "Tank 4P BWT DO", Enable :=, "Enable Delay Time" := T#0ms, "High Value Release" :=, "SHORT CIRCUIT VALUE" :=, "BROKEN WIRE VALUE" :=, "VERY LOW LEVEL VALUE (LL)" :=, "LOW LEVEL VALUE (L)" :=, "HIGH LEVEL VALUE (H)" :=, "VERY HIGH LEVEL VALUE (HH)" :=, OFFSET :=, "ALARM DELAY" := T#100ms, "Peak Value Reset" :=, "ALARM HH" =>, "ALARM H" =>, "ALARM L" =>, "ALARM LL" =>, "ALARM READING" => %DB2062.DBX372.1, "Peak Value" =>, Alarm =>, Alarm_INT =>)
   END_RUNG
   // the same network as SCL:
   "BWT 4P DO (426) ALARM"(Value := "20_TANKS_IP_DATA".RIO_04.FIRST_TANK.BWT_DO,   // "502_ALM_ANALOG"
                           "Raw Value" := "Tank 4P BWT DO",
                           "Enable Delay Time" := T#0ms,
                           "ALARM DELAY" := T#100ms,
                           "ALARM READING" => %DB2062.DBX372.1);
END_REGION

REGION Network 93: DB2062.DBX372.2 = DO426 4S
   // BTCS_WARNING_WORD_17_BIT_2
